      statAcknowledgeReqestedEStop8 : Bool;
      ESTOP1_Instance_1 : ESTOP1;
      ESTOP1_Instance_2 : ESTOP1;
      ESTOP1_Instance_3 : ESTOP1;
      ESTOP1_Instance_4 : ESTOP1;
      ESTOP1_Instance_5 : ESTOP1;
      ESTOP1_Instance_6 : ESTOP1;
      ESTOP1_Instance_7 : ESTOP1;
      ESTOP1_Instance_8 : ESTOP1;
   END_VAR
BEGIN

REGION Network 1
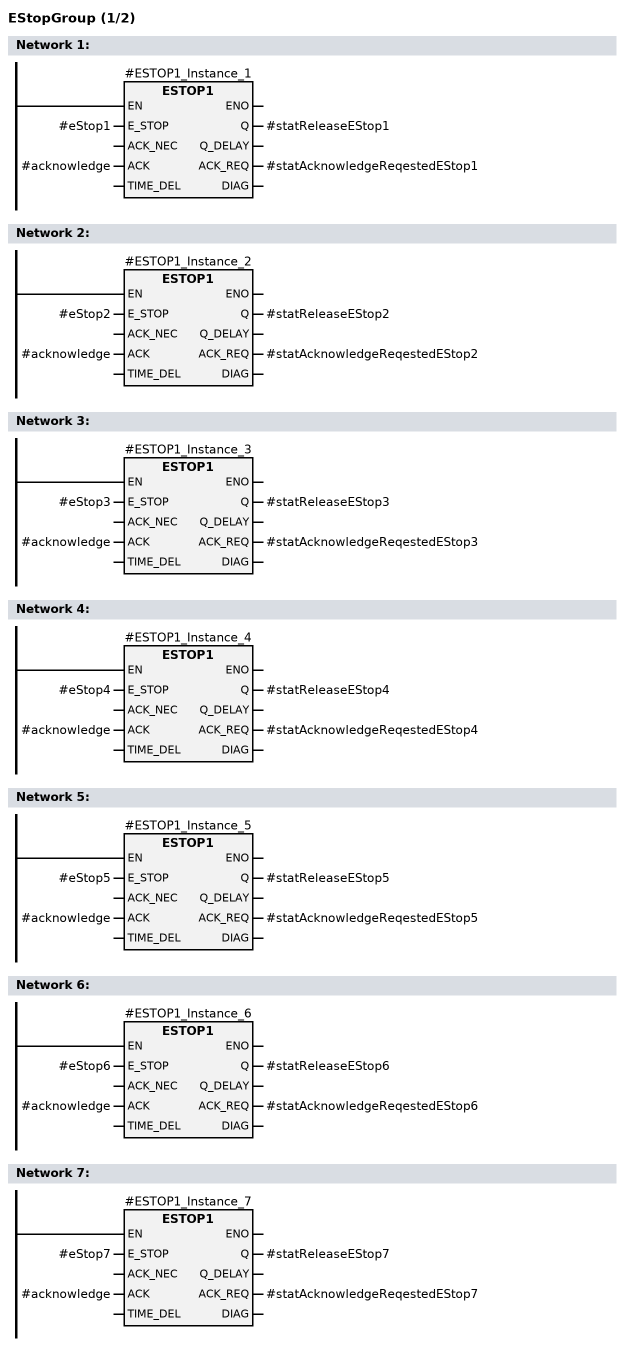
   #ESTOP1_Instance_1(E_STOP := #eStop1,   // ESTOP1
                      ACK := #acknowledge,
                      Q => #statReleaseEStop1,
                      ACK_REQ => #statAcknowledgeReqestedEStop1);
END_REGION

REGION Network 2
   #ESTOP1_Instance_2(E_STOP := #eStop2,   // ESTOP1
                      ACK := #acknowledge,
                      Q => #statReleaseEStop2,
                      ACK_REQ => #statAcknowledgeReqestedEStop2);
END_REGION

REGION Network 3
   #ESTOP1_Instance_3(E_STOP := #eStop3,   // ESTOP1
                      ACK := #acknowledge,
                      Q => #statReleaseEStop3,
                      ACK_REQ => #statAcknowledgeReqestedEStop3);
END_REGION

REGION Network 4
   #ESTOP1_Instance_4(E_STOP := #eStop4,   // ESTOP1
                      ACK := #acknowledge,
                      Q => #statReleaseEStop4,
                      ACK_REQ => #statAcknowledgeReqestedEStop4);
END_REGION

REGION Network 5
   #ESTOP1_Instance_5(E_STOP := #eStop5,   // ESTOP1
                      ACK := #acknowledge,
                      Q => #statReleaseEStop5,
                      ACK_REQ => #statAcknowledgeReqestedEStop5);
END_REGION

REGION Network 6
   #ESTOP1_Instance_6(E_STOP := #eStop6,   // ESTOP1
                      ACK := #acknowledge,
                      Q => #statReleaseEStop6,
                      ACK_REQ => #statAcknowledgeReqestedEStop6);
END_REGION

REGION Network 7
   #ESTOP1_Instance_7(E_STOP := #eStop7,   // ESTOP1
                      ACK := #acknowledge,
                      Q => #statReleaseEStop7,
                      ACK_REQ => #statAcknowledgeReqestedEStop7);
END_REGION

REGION Network 8
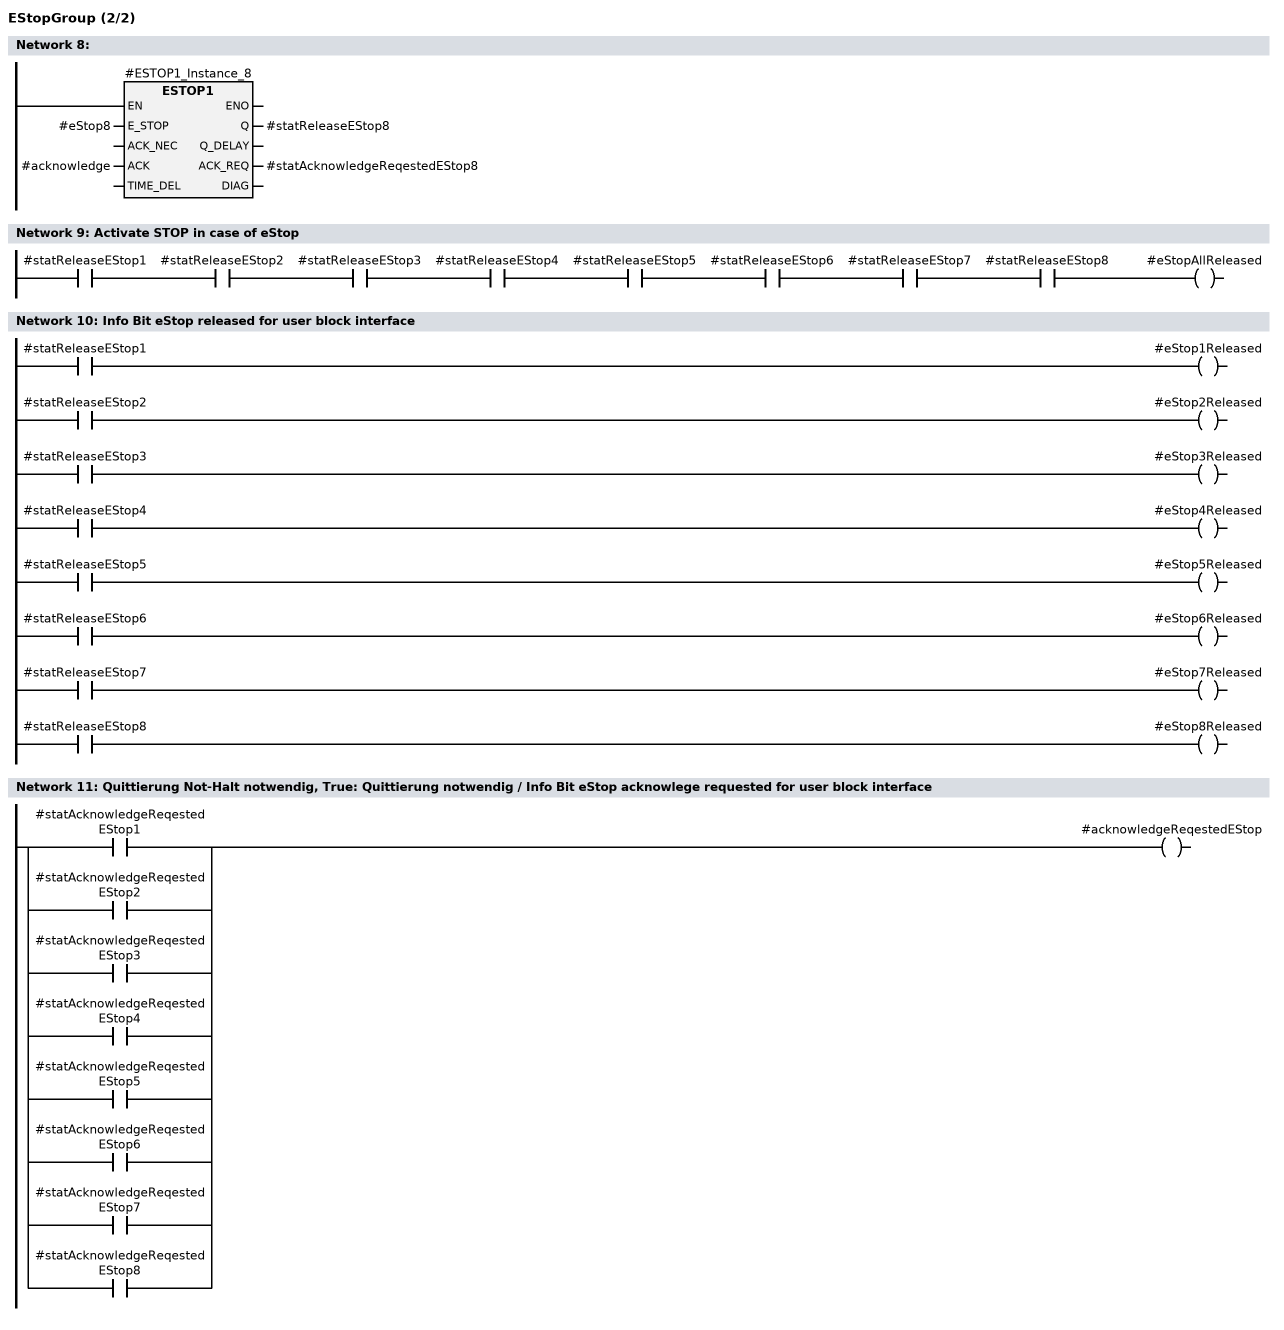
   #ESTOP1_Instance_8(E_STOP := #eStop8,   // ESTOP1
                      ACK := #acknowledge,
                      Q => #statReleaseEStop8,
                      ACK_REQ => #statAcknowledgeReqestedEStop8);
END_REGION

REGION Network 9: Activate STOP in case of eStop
   RUNG wire#powerrail
      Contact( #statReleaseEStop1 )
      Contact( #statReleaseEStop2 )
      Contact( #statReleaseEStop3 )
      Contact( #statReleaseEStop4 )
      Contact( #statReleaseEStop5 )
      Contact( #statReleaseEStop6 )
      Contact( #statReleaseEStop7 )
      Contact( #statReleaseEStop8 )
      Coil( #eStopAllReleased )
   END_RUNG
   // the same network as SCL:
   #eStopAllReleased := #statReleaseEStop1 AND #statReleaseEStop2 AND #statReleaseEStop3 AND #statReleaseEStop4 AND #statReleaseEStop5 AND #statReleaseEStop6 AND #statReleaseEStop7 AND #statReleaseEStop8;
END_REGION

REGION Network 10: Info Bit eStop released for user block interface
   RUNG wire#powerrail
      Contact( #statReleaseEStop1 )
      Coil( #eStop1Released )
   END_RUNG
   RUNG wire#powerrail
      Contact( #statReleaseEStop2 )
      Coil( #eStop2Released )
   END_RUNG
   RUNG wire#powerrail
      Contact( #statReleaseEStop3 )
      Coil( #eStop3Released )
   END_RUNG
   RUNG wire#powerrail
      Contact( #statReleaseEStop4 )
      Coil( #eStop4Released )
   END_RUNG
   RUNG wire#powerrail
      Contact( #statReleaseEStop5 )
      Coil( #eStop5Released )
   END_RUNG
   RUNG wire#powerrail
      Contact( #statReleaseEStop6 )
      Coil( #eStop6Released )
   END_RUNG
   RUNG wire#powerrail
      Contact( #statReleaseEStop7 )
      Coil( #eStop7Released )
   END_RUNG
   RUNG wire#powerrail
      Contact( #statReleaseEStop8 )
      Coil( #eStop8Released )
   END_RUNG
   // the same network as SCL:
   #eStop1Released := #statReleaseEStop1;
   #eStop2Released := #statReleaseEStop2;
   #eStop3Released := #statReleaseEStop3;
   #eStop4Released := #statReleaseEStop4;
   #eStop5Released := #statReleaseEStop5;
   #eStop6Released := #statReleaseEStop6;
   #eStop7Released := #statReleaseEStop7;
   #eStop8Released := #statReleaseEStop8;
END_REGION

REGION Network 11: Quittierung Not-Halt notwendig, True: Quittierung notwendig / Info Bit eStop acknowlege requested for user block interface
   RUNG wire#powerrail
      Contact( #statAcknowledgeReqestedEStop1 )
      wire#w1
      Coil( #acknowledgeReqestedEStop )
   END_RUNG
   RUNG wire#powerrail
      Contact( #statAcknowledgeReqestedEStop2 )
   END_RUNG wire#w1
   RUNG wire#powerrail
      Contact( #statAcknowledgeReqestedEStop3 )
   END_RUNG wire#w1
   RUNG wire#powerrail
      Contact( #statAcknowledgeReqestedEStop4 )
   END_RUNG wire#w1
   RUNG wire#powerrail
      Contact( #statAcknowledgeReqestedEStop5 )
   END_RUNG wire#w1
   RUNG wire#powerrail
      Contact( #statAcknowledgeReqestedEStop6 )
   END_RUNG wire#w1
   RUNG wire#powerrail
      Contact( #statAcknowledgeReqestedEStop7 )
   END_RUNG wire#w1
   RUNG wire#powerrail
      Contact( #statAcknowledgeReqestedEStop8 )
   END_RUNG wire#w1
   // the same network as SCL:
   #acknowledgeReqestedEStop := #statAcknowledgeReqestedEStop1 OR #statAcknowledgeReqestedEStop2 OR #statAcknowledgeReqestedEStop3 OR #statAcknowledgeReqestedEStop4 OR #statAcknowledgeReqestedEStop5 OR #statAcknowledgeReqestedEStop6 OR #statAcknowledgeReqestedEStop7 OR #statAcknowledgeReqestedEStop8;
END_REGION
END_FUNCTION_BLOCK

FUNCTION_BLOCK "LightCurtainGroup"   // FB12, F_LAD
{ S7_Optimized_Access := 'TRUE' }
VERSION : 0.1
   VAR_INPUT
      acknowledge : Bool;   // Acknowledge / Quittierung, Positive Flanke notwendig, NO / Acknowledge, positive signal edge, NO
      selAccZone : Bool;
      entryButtonZone1 : Bool;   // Entry button – Zone 1 (LC 1-6)
      entryButtonZone2 : Bool;   // Entry button – Zone 2 (LC 1, 3, 6)
      entryButtonZone3 : Bool;   // Entry button – Zone 3 (LC 2, 4, 5)
      robotInZone2 : Bool;
      robotInZone3 : Bool;
      lc1Ossd1 : Bool;
      lc1Ossd2 : Bool;
      lc2Ossd1 : Bool;
      lc2Ossd2 : Bool;
      lc3Ossd1 : Bool;
      lc3Ossd2 : Bool;
      lc4Ossd1 : Bool;
      lc4Ossd2 : Bool;
      lc5Ossd1 : Bool;
      lc5Ossd2 : Bool;
      lc6Ossd1 : Bool;
      lc6Ossd2 : Bool;
   END_VAR
   VAR_OUTPUT
      lcAllFree : Bool;   // All light curtains ready
      lc1Free : Bool;   // Light curtain 1 ready
      lc2Free : Bool;
      lc3Free : Bool;   // Light curtain 3 ready
      lc4Free : Bool;
      lc5Free : Bool;
      lc6Free : Bool;   // Light curtain 6 ready
      accessReqZ2 : Bool;
      accessReqZ3 : Bool;
      zone1AccessGranted : Bool;
      zone2AccessGranted : Bool;
      zone3AccessGranted : Bool;
   END_VAR
   VAR
      EV1oo2DI_Instance_1 : EV1oo2DI;
      EV1oo2DI_Instance_2 : EV1oo2DI;
      EV1oo2DI_Instance_3 : EV1oo2DI;
      MUT_P_Instance_1 : MUT_P;
      accZ2Ok : Bool;
      accZ3Ok : Bool;
      lcZone2Free : Bool;
      lcZone3Free : Bool;
      EV1oo2DI_Instance_4 : EV1oo2DI;
      EV1oo2DI_Instance_5 : EV1oo2DI;
      EV1oo2DI_Instance_6 : EV1oo2DI;
   END_VAR
BEGIN

REGION Network 1
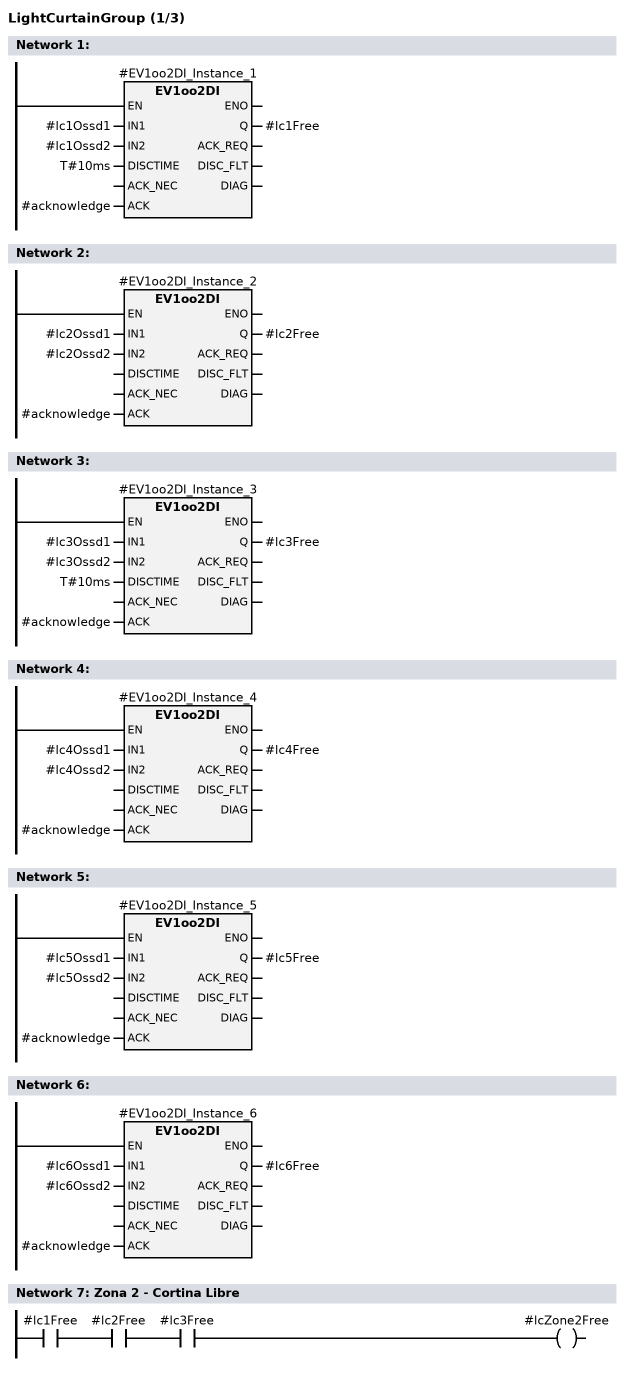
   #EV1oo2DI_Instance_1(IN1 := #lc1Ossd1,   // EV1oo2DI
                        IN2 := #lc1Ossd2,
                        DISCTIME := T#10ms,
                        ACK := #acknowledge,
                        Q => #lc1Free);
END_REGION

REGION Network 2
   #EV1oo2DI_Instance_2(IN1 := #lc2Ossd1, IN2 := #lc2Ossd2, ACK := #acknowledge, Q => #lc2Free);   // EV1oo2DI
END_REGION

REGION Network 3
   #EV1oo2DI_Instance_3(IN1 := #lc3Ossd1,   // EV1oo2DI
                        IN2 := #lc3Ossd2,
                        DISCTIME := T#10ms,
                        ACK := #acknowledge,
                        Q => #lc3Free);
END_REGION

REGION Network 4
   #EV1oo2DI_Instance_4(IN1 := #lc4Ossd1, IN2 := #lc4Ossd2, ACK := #acknowledge, Q => #lc4Free);   // EV1oo2DI
END_REGION

REGION Network 5
   #EV1oo2DI_Instance_5(IN1 := #lc5Ossd1, IN2 := #lc5Ossd2, ACK := #acknowledge, Q => #lc5Free);   // EV1oo2DI
END_REGION

REGION Network 6
   #EV1oo2DI_Instance_6(IN1 := #lc6Ossd1, IN2 := #lc6Ossd2, ACK := #acknowledge, Q => #lc6Free);   // EV1oo2DI
END_REGION

REGION Network 7: Zona 2 - Cortina Libre
   RUNG wire#powerrail
      Contact( #lc1Free )
      Contact( #lc2Free )
      Contact( #lc3Free )
      Coil( #lcZone2Free )
   END_RUNG
   // the same network as SCL:
   #lcZone2Free := #lc1Free AND #lc2Free AND #lc3Free;
END_REGION

REGION Network 8: Zona 3 - Cortina Libre
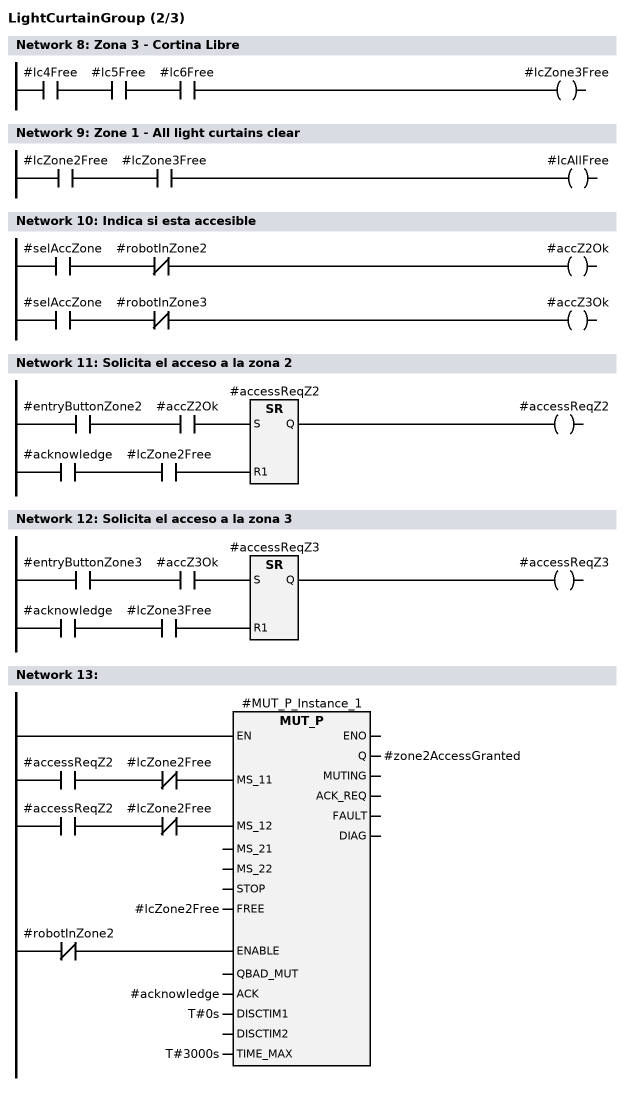
   RUNG wire#powerrail
      Contact( #lc4Free )
      Contact( #lc5Free )
      Contact( #lc6Free )
      Coil( #lcZone3Free )
   END_RUNG
   // the same network as SCL:
   #lcZone3Free := #lc4Free AND #lc5Free AND #lc6Free;
END_REGION

REGION Network 9: Zone 1 - All light curtains clear
   RUNG wire#powerrail
      Contact( #lcZone2Free )
      Contact( #lcZone3Free )
      Coil( #lcAllFree )
   END_RUNG
   // the same network as SCL:
   #lcAllFree := #lcZone2Free AND #lcZone3Free;
END_REGION

REGION Network 10: Indica si esta accesible
   RUNG wire#powerrail
      Contact( #selAccZone )
      I_Contact( #robotInZone2 )
      Coil( #accZ2Ok )
   END_RUNG
   RUNG wire#powerrail
      Contact( #selAccZone )
      I_Contact( #robotInZone3 )
      Coil( #accZ3Ok )
   END_RUNG
   // the same network as SCL:
   #accZ2Ok := #selAccZone AND NOT #robotInZone2;
   #accZ3Ok := #selAccZone AND NOT #robotInZone3;
END_REGION

REGION Network 11: Solicita el acceso a la zona 2
   RUNG wire#powerrail
      Contact( #entryButtonZone2 )
      Contact( #accZ2Ok )
      S_SR(operand := #accessReqZ2, r1 := wire#w1)
      Coil( #accessReqZ2 )
   END_RUNG
   RUNG wire#powerrail
      Contact( #acknowledge )
      Contact( #lcZone2Free )
   END_RUNG wire#w1
   // the same network as SCL:
   IF #entryButtonZone2 AND #accZ2Ok THEN
       #accessReqZ2 := TRUE;   // SR flip-flop
   END_IF;
   IF #acknowledge AND #lcZone2Free THEN #accessReqZ2 := FALSE; END_IF;
   #accessReqZ2 := #accessReqZ2;
END_REGION

REGION Network 12: Solicita el acceso a la zona 3
   RUNG wire#powerrail
      Contact( #entryButtonZone3 )
      Contact( #accZ3Ok )
      S_SR(operand := #accessReqZ3, r1 := wire#w1)
      Coil( #accessReqZ3 )
   END_RUNG
   RUNG wire#powerrail
      Contact( #acknowledge )
      Contact( #lcZone3Free )
   END_RUNG wire#w1
   // the same network as SCL:
   IF #entryButtonZone3 AND #accZ3Ok THEN
       #accessReqZ3 := TRUE;   // SR flip-flop
   END_IF;
   IF #acknowledge AND #lcZone3Free THEN #accessReqZ3 := FALSE; END_IF;
   #accessReqZ3 := #accessReqZ3;
END_REGION

REGION Network 13
   #MUT_P_Instance_1(MS_11 := #accessReqZ2 AND NOT #lcZone2Free,   // MUT_P
                     MS_12 := #accessReqZ2 AND NOT #lcZone2Free,
                     FREE := #lcZone2Free,
                     ENABLE := NOT #robotInZone2,
                     ACK := #acknowledge,
                     DISCTIM1 := T#0s,
                     TIME_MAX := T#3000s,
                     Q => #zone2AccessGranted);
END_REGION

REGION Network 14
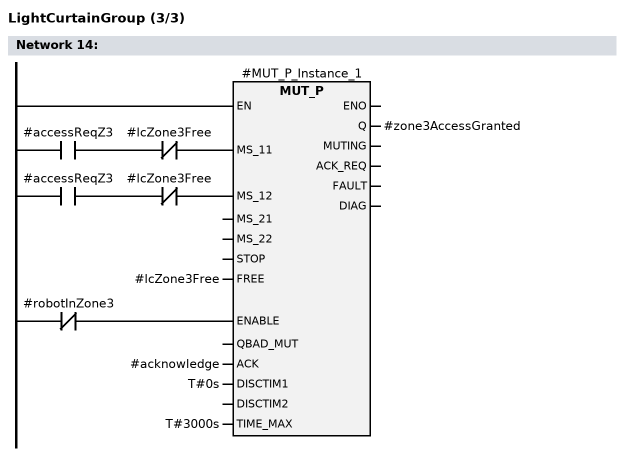
   #MUT_P_Instance_1(MS_11 := #accessReqZ3 AND NOT #lcZone3Free,   // MUT_P
                     MS_12 := #accessReqZ3 AND NOT #lcZone3Free,
                     FREE := #lcZone3Free,
                     ENABLE := NOT #robotInZone3,
                     ACK := #acknowledge,
                     DISCTIM1 := T#0s,
                     TIME_MAX := T#3000s,
                     Q => #zone3AccessGranted);
END_REGION
END_FUNCTION_BLOCK

FUNCTION_BLOCK "SafetyDoor"   // FB13, F_FBD
{ S7_Optimized_Access := 'TRUE' }
VERSION : 0.1
   VAR_OUTPUT
      SAF_DOOR_CLSD_RDY : Bool;   // Safety door closed & locked – ready
   END_VAR
   VAR
      SFDOOR_Instance_1 : SFDOOR;
   END_VAR
BEGIN

REGION Network 1
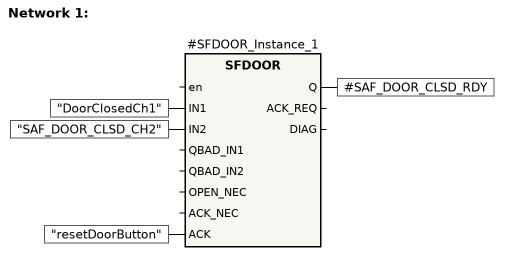
   #SFDOOR_Instance_1(IN1 := "DoorClosedCh1",   // SFDOOR
                      IN2 := "SAF_DOOR_CLSD_CH2",
                      ACK := "resetDoorButton",
                      Q => #SAF_DOOR_CLSD_RDY);
END_REGION
END_FUNCTION_BLOCK

(* ===== HMI "HMI_RT_1" =====
system functions are stored by id; their names below are inferred from use
connection "HMI_Connection_1": ETHERNET, SMART_S7_1200_OMS

HMI tags "Default tag table"
   "Tag_ScreenNumber" : UInt, internal

Template "Template_1" 1280x800
   Button "Exit" at 1182,752 size 67x47; TextOff 'Exit'; PictureOff "ExitRuntime_KTP1200_Basic_PN_TR"; PictureOn "ExitRuntime_KTP1200_Basic_PN_TR"
      on Release: StopRuntime(0)
   Button "Template_Button" at 1054,752 size 67x47; TextOff 'Text'
   Button "Template_Button_1" at 926,752 size 67x47; TextOff 'Text'
   Button "Template_Button_2" at 798,752 size 67x47; TextOff 'Text'
   Button "Template_Button_3" at 670,752 size 67x47; TextOff 'Text'
   Button "Template_Button_4" at 542,752 size 67x47; TextOff 'Text'
   Button "Template_Button_5" at 414,752 size 67x47; TextOff 'Text'
   Button "Template_Button_6" at 286,752 size 67x47; TextOff 'Text'
   Button "Alarms" at 158,752 size 67x47; TextOff 'Alarms'; PictureOff "AlarmDisplay_KTP1200_Basic_PN_TR"; PictureOn "AlarmDisplay_KTP1200_Basic_PN_TR"
      on Release: function_ef3f5d25("Alarm window_Unacknowledged", -1)
   Button "Start screen" at 30,752 size 67x47; TextOff 'Start screen'; PictureOff "NavigateHome_KTP1200_Basic_PN_TR"; PictureOn "NavigateHome_KTP1200_Basic_PN_TR"
      on Release: ActivateScreen("Root screen", 0)
   SymbolicIOField "Symbolic_IO_Field_Screen" at 87,9 size 1086x30; TextOff '0'; TextOn '1'; TextList "TextList_ScreenNames"
      ProcessValue <- "Tag_ScreenNumber"
      on Change: ActivateScreenByNumber("Tag_ScreenNumber", 0)
   DateTimeField "HmiScreenItemData" at 1175,24 size 105x24
   DateTimeField "HmiScreenItemData_1" at 1175,0 size 105x24
   GraphicView "Logo" at 0,0 size 85x48; Picture "Logo of HMI_1"

screen "Root screen" 1280x800, template "Template_1"
   on GenerateScreen: SetTag("Tag_ScreenNumber", 1)
   TextField "HmiScreenItemData_1" at 128,384 size 1024x27; Text 'Welcome to HMI_1 (KTP1200 Basic+ PN)!'
   Button "HmiScreenItemData" at 36,84 size 159x47; TextOff 'Screen_Prueba'; PictureOff "Navigates to Screen_Prueba for KTP1200 Basic+ PN 17.0.0.0"; PictureOn "Navigates to Screen_Prueba for KTP1200 Basic+ PN 17.0.0.0"
      on Release: ActivateScreen("Screen_Prueba", 0)
   Button "HmiScreenItemData_2" at 36,143 size 159x47; TextOff 'System screens'; PictureOff "Navigates to System screens for KTP1200 Basic+ PN 17.0.0.0"; PictureOn "Navigates to System screens for KTP1200 Basic+ PN 17.0.0.0"
      on Release: ActivateScreen("System screens", 0)

screen "Screen_Prueba" 1280x800, template "Template_1"
   on GenerateScreen: SetTag("Tag_ScreenNumber", 2)
   TextField "HmiScreenItemData" at 128,384 size 1024x27; Text 'Screen_Prueba'
   Button "Back" at 1,49 size 159x47; TextOff 'Back'
      on Release: ActivateScreen("Root screen", 0)

screen "System screens" 1280x800, template "Template_1"
   on GenerateScreen: SetTag("Tag_ScreenNumber", 3)
   Button "Back" at 1,49 size 159x47; TextOff 'Back'
      on Release: ActivateScreen("Root screen", 0)
   Button "HmiScreenItemData" at 36,143 size 159x47; TextOff 'SIMATIC PLC system diagnos...'; PictureOff "Navigates to SIMATIC PLC system diagnostics for KTP1200 Basic+ PN 17.0.0.0"; PictureOn "Navigates to SIMATIC PLC system diagnostics for KTP1200 Basic+ PN 17.0.0.0"
      on Release: ActivateScreen("SIMATIC PLC system diagnostics", 0)
   Button "HmiScreenItemData_1" at 36,202 size 159x47; TextOff 'Project information'; PictureOff "Navigates to Project information for KTP1200 Basic+ PN 17.0.0.0"; PictureOn "Navigates to Project information for KTP1200 Basic+ PN 17.0.0.0"
      on Release: ActivateScreen("Project information", 0)
   Button "HmiScreenItemData_2" at 36,261 size 159x47; TextOff 'User administration'; PictureOff "Navigates to User administration for KTP1200 Basic+ PN 17.0.0.0"; PictureOn "Navigates to User administration for KTP1200 Basic+ PN 17.0.0.0"
      on Release: ActivateScreen("User administration", 0)
   Button "HmiScreenItemData_3" at 36,320 size 159x47; TextOff 'System information'; PictureOff "Navigates to System information for KTP1200 Basic+ PN 17.0.0.0"; PictureOn "Navigates to System information for KTP1200 Basic+ PN 17.0.0.0"
      on Release: ActivateScreen("System information", 0)
   Button "HmiScreenItemData_4" at 36,379 size 159x47; TextOff 'Different jobs'; PictureOff "Navigates to Different jobs for KTP1200 Basic+ PN 17.0.0.0"; PictureOn "Navigates to Different jobs for KTP1200 Basic+ PN 17.0.0.0"
      on Release: ActivateScreen("Different jobs", 0)

screen "SIMATIC PLC system diagnostics" 1280x800, template "Template_1"
   on GenerateScreen: SetTag("Tag_ScreenNumber", 4)
   SysDiagControl "HmiScreenItemData" at 1,97 size 1276x647
   Button "Back" at 1,49 size 159x47; TextOff 'Back'
      on Release: ActivateScreen("System screens", 0)

screen "Project information" 1280x800, template "Template_1"
   on GenerateScreen: SetTag("Tag_ScreenNumber", 5)
   TextField "HmiScreenItemData" at 35,99 size 171x28; Text 'Project name:'
   TextField "HmiScreenItemData_1" at 241,99 size 1004x28; Text 'HEAT-1-CADIZ-V5'
   TextField "HmiScreenItemData_2" at 35,129 size 171x28; Text 'Created on:'
   TextField "HmiScreenItemData_3" at 241,129 size 1004x28; Text '4/3/2025 12:55:11 PM'
   TextField "HmiScreenItemData_4" at 35,159 size 171x28; Text 'Author:'
   TextField "HmiScreenItemData_5" at 241,159 size 1004x28; Text 'User'
   TextField "HmiScreenItemData_6" at 35,189 size 171x28; Text 'Description:'
   TextField "HmiScreenItemData_7" at 241,189 size 1004x28; Text '(not configured)'
   Button "Back" at 1,49 size 159x47; TextOff 'Back'
      on Release: ActivateScreen("System screens", 0)

screen "User administration" 1280x800, template "Template_1"
   on GenerateScreen: SetTag("Tag_ScreenNumber", 6)
   UserView "HmiScreenItemData" at 1,97 size 1276x647
   Button "Back" at 1,49 size 159x47; TextOff 'Back'
      on Release: ActivateScreen("System screens", 0)

screen "System information" 1280x800, template "Template_1"
   on GenerateScreen: SetTag("Tag_ScreenNumber", 7)
   TextField "HmiScreenItemData" at 35,99 size 171x28; Text 'HMI device type:'
   TextField "HmiScreenItemData_1" at 241,99 size 1004x28; Text 'KTP1200 Basic+ PN 17.0.0.0'
   TextField "HmiScreenItemData_2" at 35,129 size 171x28; Text 'Connection:'
   TextField "HmiScreenItemData_3" at 241,129 size 1004x28; Text 'PROFINET (X1)'
   TextField "HmiScreenItemData_4" at 35,159 size 171x28; Text 'PLC:'
   TextField "HmiScreenItemData_5" at 241,159 size 1004x28; Text 'SIMATIC S7 1200'
   Button "Back" at 1,49 size 159x47; TextOff 'Back'
      on Release: ActivateScreen("System screens", 0)

screen "Different jobs" 1280x800, template "Template_1"
   on GenerateScreen: SetTag("Tag_ScreenNumber", 8)
   Button "Online" at 36,143 size 159x47; TextOff 'Online'
      on Release: function_bb44b551(0)
   Button "Offline" at 36,202 size 159x47; TextOff 'Offline'
      on Release: function_bb44b551(1)
   Button "Transfer" at 36,261 size 159x47; TextOff 'Transfer'
      on Release: function_bb44b551(2)
   Button "Toggle language" at 36,320 size 159x47; TextOff 'Toggle language'
      on Release: function_fb9197e8(-1)
   Button "Stop Runtime" at 36,379 size 159x47; TextOff 'Stop Runtime'
      on Release: StopRuntime(0)
   Button "Back" at 1,49 size 159x47; TextOff 'Back'
      on Release: ActivateScreen("System screens", 0)
*)